DATA_BLOCK "DB_SDC_TS_PARAMETER_4"   // DB3707
{ S7_Optimized_Access := 'FALSE' }
AUTHOR : FFM
FAMILY : SDC
NAME : SECT_DEF
VERSION : 1.0
   VAR
      HEADER : Struct   // Struktur für Datenheader // nicht verschieben
         DB_NR : Int := 3707;   // DB Nummer
         MIN_NR_SEK : Int := 301;   // Niedrigste SEK Nummer im DB
         MAX_NR_SEK : Int := 400;   // Höchste SEK Nummer im DB
         START_DAT : Int := 20;   // Startadresse der SEK im DB
         LAENGE_SEK_DATA : Int := 260;   // Länge SEK Data
         ANZ_PROFIL : Int := 10;   // Number of Profiles
         OFFEST_PROFIL : Int := 40;   // Offestadresse der Profilparameter im TS-Parameterdatensatz
         LAENGE_PROFIL_DATA : Int := 22;   // Länge SEK Data
         Res160 : Int := 0;   // Reserve
         Res : Int := 0;   // Reserve
      END_STRUCT;
      TS : Array[301..400] of "UDT_SDC_TS_PARAMETER";
   END_VAR
BEGIN
   TS[301].ALLG.SEK_NEXT_1 := 0;
   TS[301].ALLG.SEK_NEXT_2 := 0;
   TS[301].ALLG.Spare[4] := 16#00;
   TS[301].ALLG.Spare[5] := 16#00;
   TS[301].ALLG.POS.Start_1 := 0;
   TS[301].ALLG.POS.End_1 := 0;
   TS[301].ALLG.POS.Start_2 := 0;
   TS[301].ALLG.POS.End_2 := 0;
   TS[301].ALLG.POS.Actionpoint_1 := 0;
   TS[301].ALLG.POS.Actionpoint_2 := 0;
   TS[301].ALLG.FLAGS.DIST_VAL[0] := TRUE;
   TS[301].ALLG.FLAGS.DIST_VAL[1] := FALSE;
   TS[301].ALLG.FLAGS.DIST_VAL[2] := FALSE;
   TS[301].ALLG.FLAGS.DIST_VAL[3] := FALSE;
   TS[301].ALLG.FLAGS.DIST_VAL[4] := FALSE;
   TS[301].ALLG.FLAGS.DIST_VAL[5] := FALSE;
   TS[301].ALLG.FLAGS.DIST_VAL[6] := FALSE;
   TS[301].ALLG.FLAGS.DIST_VAL[7] := FALSE;
   TS[301].ALLG.FLAGS.DIST_VAL[8] := FALSE;
   TS[301].ALLG.FLAGS.DIST_VAL[9] := FALSE;
   TS[301].ALLG.FLAGS.DIST_VAL[10] := FALSE;
   TS[301].ALLG.FLAGS.DIST_VAL[11] := FALSE;
   TS[301].ALLG.FLAGS.DIST_VAL[12] := FALSE;
   TS[301].ALLG.FLAGS.DIST_VAL[13] := FALSE;
   TS[301].ALLG.FLAGS.DIST_VAL[14] := FALSE;
   TS[301].ALLG.FLAGS.DIST_VAL[15] := FALSE;
   TS[301].ALLG.FLAGS.one_profile := FALSE;
   TS[301].ALLG.FLAGS.BLIND := FALSE;
   TS[301].ALLG.FLAGS.NO_DIST_CONT := FALSE;
   TS[301].ALLG.FLAGS.SYNCH_AREA := FALSE;
   TS[301].ALLG.FLAGS.bit24 := FALSE;
   TS[301].ALLG.FLAGS.bit25 := FALSE;
   TS[301].ALLG.FLAGS.bit26 := FALSE;
   TS[301].ALLG.FLAGS.bit27 := FALSE;
   TS[301].ALLG.FLAGS.EN_HOIST := FALSE;
   TS[301].ALLG.FLAGS.D_RESET_AFTER := FALSE;
   TS[301].ALLG.FLAGS.D_PULK := FALSE;
   TS[301].ALLG.FLAGS.bit33 := FALSE;
   TS[301].ALLG.FLAGS.bit34 := FALSE;
   TS[301].ALLG.FLAGS.bit35 := FALSE;
   TS[301].ALLG.FLAGS.bit36 := FALSE;
   TS[301].ALLG.FLAGS.Deutronic_ON := FALSE;
   TS[301].ALLG.Stop_Position := 0;
   TS[301].ALLG.Drive_speed_1 := 0;
   TS[301].ALLG.Drive_speed_2 := 0;
   TS[301].PROFIL[1].Hoist_Pos_start := 0;
   TS[301].PROFIL[1].Height := 2651;
   TS[301].PROFIL[1].Hoist_speed := 2000;
   TS[301].PROFIL[1].Hoist_offset_1 := 0;
   TS[301].PROFIL[1].Hoist_offset_2 := 0;
   TS[301].PROFIL[1].Hoist_offset_3 := 0;
   TS[301].PROFIL[1].Hoist_offset_4 := 0;
   TS[301].PROFIL[1].Hoist_Start_offset_1 := 0;
   TS[301].PROFIL[1].Hoist_Start_offset_2 := 0;
   TS[301].PROFIL[1].Hoist_Start_offset_3 := 0;
   TS[301].PROFIL[1].Hoist_Start_offset_4 := 0;
   TS[301].PROFIL[2].Hoist_Pos_start := 0;
   TS[301].PROFIL[2].Height := 2651;
   TS[301].PROFIL[2].Hoist_speed := 2000;
   TS[301].PROFIL[2].Hoist_offset_1 := 0;
   TS[301].PROFIL[2].Hoist_offset_2 := 0;
   TS[301].PROFIL[2].Hoist_offset_3 := 0;
   TS[301].PROFIL[2].Hoist_offset_4 := 0;
   TS[301].PROFIL[2].Hoist_Start_offset_1 := 0;
   TS[301].PROFIL[2].Hoist_Start_offset_2 := 0;
   TS[301].PROFIL[2].Hoist_Start_offset_3 := 0;
   TS[301].PROFIL[2].Hoist_Start_offset_4 := 0;
   TS[301].PROFIL[3].Hoist_Pos_start := 0;
   TS[301].PROFIL[3].Height := 2651;
   TS[301].PROFIL[3].Hoist_speed := 2000;
   TS[301].PROFIL[3].Hoist_offset_1 := 0;
   TS[301].PROFIL[3].Hoist_offset_2 := 0;
   TS[301].PROFIL[3].Hoist_offset_3 := 0;
   TS[301].PROFIL[3].Hoist_offset_4 := 0;
   TS[301].PROFIL[3].Hoist_Start_offset_1 := 0;
   TS[301].PROFIL[3].Hoist_Start_offset_2 := 0;
   TS[301].PROFIL[3].Hoist_Start_offset_3 := 0;
   TS[301].PROFIL[3].Hoist_Start_offset_4 := 0;
   TS[301].PROFIL[4].Hoist_Pos_start := 0;
   TS[301].PROFIL[4].Height := 2651;
   TS[301].PROFIL[4].Hoist_speed := 2000;
   TS[301].PROFIL[4].Hoist_offset_1 := 0;
   TS[301].PROFIL[4].Hoist_offset_2 := 0;
   TS[301].PROFIL[4].Hoist_offset_3 := 0;
   TS[301].PROFIL[4].Hoist_offset_4 := 0;
   TS[301].PROFIL[4].Hoist_Start_offset_1 := 0;
   TS[301].PROFIL[4].Hoist_Start_offset_2 := 0;
   TS[301].PROFIL[4].Hoist_Start_offset_3 := 0;
   TS[301].PROFIL[4].Hoist_Start_offset_4 := 0;
   TS[301].PROFIL[5].Hoist_Pos_start := 0;
   TS[301].PROFIL[5].Height := 2651;
   TS[301].PROFIL[5].Hoist_speed := 2000;
   TS[301].PROFIL[5].Hoist_offset_1 := 0;
   TS[301].PROFIL[5].Hoist_offset_2 := 0;
   TS[301].PROFIL[5].Hoist_offset_3 := 0;
   TS[301].PROFIL[5].Hoist_offset_4 := 0;
   TS[301].PROFIL[5].Hoist_Start_offset_1 := 0;
   TS[301].PROFIL[5].Hoist_Start_offset_2 := 0;
   TS[301].PROFIL[5].Hoist_Start_offset_3 := 0;
   TS[301].PROFIL[5].Hoist_Start_offset_4 := 0;
   TS[301].PROFIL[6].Hoist_Pos_start := 0;
   TS[301].PROFIL[6].Height := 2651;
   TS[301].PROFIL[6].Hoist_speed := 2000;
   TS[301].PROFIL[6].Hoist_offset_1 := 0;
   TS[301].PROFIL[6].Hoist_offset_2 := 0;
   TS[301].PROFIL[6].Hoist_offset_3 := 0;
   TS[301].PROFIL[6].Hoist_offset_4 := 0;
   TS[301].PROFIL[6].Hoist_Start_offset_1 := 0;
   TS[301].PROFIL[6].Hoist_Start_offset_2 := 0;
   TS[301].PROFIL[6].Hoist_Start_offset_3 := 0;
   TS[301].PROFIL[6].Hoist_Start_offset_4 := 0;
   TS[301].PROFIL[7].Hoist_Pos_start := 0;
   TS[301].PROFIL[7].Height := 2651;
   TS[301].PROFIL[7].Hoist_speed := 2000;
   TS[301].PROFIL[7].Hoist_offset_1 := 0;
   TS[301].PROFIL[7].Hoist_offset_2 := 0;
   TS[301].PROFIL[7].Hoist_offset_3 := 0;
   TS[301].PROFIL[7].Hoist_offset_4 := 0;
   TS[301].PROFIL[7].Hoist_Start_offset_1 := 0;
   TS[301].PROFIL[7].Hoist_Start_offset_2 := 0;
   TS[301].PROFIL[7].Hoist_Start_offset_3 := 0;
   TS[301].PROFIL[7].Hoist_Start_offset_4 := 0;
   TS[301].PROFIL[8].Hoist_Pos_start := 0;
   TS[301].PROFIL[8].Height := 2651;
   TS[301].PROFIL[8].Hoist_speed := 2000;
   TS[301].PROFIL[8].Hoist_offset_1 := 0;
   TS[301].PROFIL[8].Hoist_offset_2 := 0;
   TS[301].PROFIL[8].Hoist_offset_3 := 0;
   TS[301].PROFIL[8].Hoist_offset_4 := 0;
   TS[301].PROFIL[8].Hoist_Start_offset_1 := 0;
   TS[301].PROFIL[8].Hoist_Start_offset_2 := 0;
   TS[301].PROFIL[8].Hoist_Start_offset_3 := 0;
   TS[301].PROFIL[8].Hoist_Start_offset_4 := 0;
   TS[301].PROFIL[9].Hoist_Pos_start := 0;
   TS[301].PROFIL[9].Height := 2651;
   TS[301].PROFIL[9].Hoist_speed := 2000;
   TS[301].PROFIL[9].Hoist_offset_1 := 0;
   TS[301].PROFIL[9].Hoist_offset_2 := 0;
   TS[301].PROFIL[9].Hoist_offset_3 := 0;
   TS[301].PROFIL[9].Hoist_offset_4 := 0;
   TS[301].PROFIL[9].Hoist_Start_offset_1 := 0;
   TS[301].PROFIL[9].Hoist_Start_offset_2 := 0;
   TS[301].PROFIL[9].Hoist_Start_offset_3 := 0;
   TS[301].PROFIL[9].Hoist_Start_offset_4 := 0;
   TS[301].PROFIL[10].Hoist_Pos_start := 0;
   TS[301].PROFIL[10].Height := 2651;
   TS[301].PROFIL[10].Hoist_speed := 2000;
   TS[301].PROFIL[10].Hoist_offset_1 := 0;
   TS[301].PROFIL[10].Hoist_offset_2 := 0;
   TS[301].PROFIL[10].Hoist_offset_3 := 0;
   TS[301].PROFIL[10].Hoist_offset_4 := 0;
   TS[301].PROFIL[10].Hoist_Start_offset_1 := 0;
   TS[301].PROFIL[10].Hoist_Start_offset_2 := 0;
   TS[301].PROFIL[10].Hoist_Start_offset_3 := 0;
   TS[301].PROFIL[10].Hoist_Start_offset_4 := 0;
   TS[302].ALLG.SEK_NEXT_1 := 0;
   TS[302].ALLG.SEK_NEXT_2 := 0;
   TS[302].ALLG.Spare[4] := 16#00;
   TS[302].ALLG.Spare[5] := 16#00;
   TS[302].ALLG.POS.Start_1 := 0;
   TS[302].ALLG.POS.End_1 := 0;
   TS[302].ALLG.POS.Start_2 := 0;
   TS[302].ALLG.POS.End_2 := 0;
   TS[302].ALLG.POS.Actionpoint_1 := 0;
   TS[302].ALLG.POS.Actionpoint_2 := 0;
   TS[302].ALLG.FLAGS.DIST_VAL[0] := TRUE;
   TS[302].ALLG.FLAGS.DIST_VAL[1] := FALSE;
   TS[302].ALLG.FLAGS.DIST_VAL[2] := FALSE;
   TS[302].ALLG.FLAGS.DIST_VAL[3] := FALSE;
   TS[302].ALLG.FLAGS.DIST_VAL[4] := FALSE;
   TS[302].ALLG.FLAGS.DIST_VAL[5] := FALSE;
   TS[302].ALLG.FLAGS.DIST_VAL[6] := FALSE;
   TS[302].ALLG.FLAGS.DIST_VAL[7] := FALSE;
   TS[302].ALLG.FLAGS.DIST_VAL[8] := FALSE;
   TS[302].ALLG.FLAGS.DIST_VAL[9] := FALSE;
   TS[302].ALLG.FLAGS.DIST_VAL[10] := FALSE;
   TS[302].ALLG.FLAGS.DIST_VAL[11] := FALSE;
   TS[302].ALLG.FLAGS.DIST_VAL[12] := FALSE;
   TS[302].ALLG.FLAGS.DIST_VAL[13] := FALSE;
   TS[302].ALLG.FLAGS.DIST_VAL[14] := FALSE;
   TS[302].ALLG.FLAGS.DIST_VAL[15] := FALSE;
   TS[302].ALLG.FLAGS.one_profile := FALSE;
   TS[302].ALLG.FLAGS.BLIND := FALSE;
   TS[302].ALLG.FLAGS.NO_DIST_CONT := FALSE;
   TS[302].ALLG.FLAGS.SYNCH_AREA := FALSE;
   TS[302].ALLG.FLAGS.bit24 := FALSE;
   TS[302].ALLG.FLAGS.bit25 := FALSE;
   TS[302].ALLG.FLAGS.bit26 := FALSE;
   TS[302].ALLG.FLAGS.bit27 := FALSE;
   TS[302].ALLG.FLAGS.EN_HOIST := FALSE;
   TS[302].ALLG.FLAGS.D_RESET_AFTER := FALSE;
   TS[302].ALLG.FLAGS.D_PULK := FALSE;
   TS[302].ALLG.FLAGS.bit33 := FALSE;
   TS[302].ALLG.FLAGS.bit34 := FALSE;
   TS[302].ALLG.FLAGS.bit35 := FALSE;
   TS[302].ALLG.FLAGS.bit36 := FALSE;
   TS[302].ALLG.FLAGS.Deutronic_ON := FALSE;
   TS[302].ALLG.Stop_Position := 0;
   TS[302].ALLG.Drive_speed_1 := 0;
   TS[302].ALLG.Drive_speed_2 := 0;
   // 15300 more start values not shown
END_DATA_BLOCK

DATA_BLOCK "DB_SDC_TS_PARAMETER_5"   // DB3708
{ S7_Optimized_Access := 'FALSE' }
AUTHOR : FFM
FAMILY : SDC
NAME : SECT_DEF
VERSION : 1.0
   VAR
      HEADER : Struct   // Struktur für Datenheader // nicht verschieben
         DB_NR : Int := 3708;   // DB Nummer
         MIN_NR_SEK : Int := 401;   // Niedrigste SEK Nummer im DB
         MAX_NR_SEK : Int := 500;   // Höchste SEK Nummer im DB
         START_DAT : Int := 20;   // Startadresse der SEK im DB
         LAENGE_SEK_DATA : Int := 260;   // Länge SEK Data
         ANZ_PROFIL : Int := 10;   // Number of Profiles
         OFFEST_PROFIL : Int := 40;   // Offestadresse der Profilparameter im TS-Parameterdatensatz
         LAENGE_PROFIL_DATA : Int := 22;   // Länge SEK Data
         Res160 : Int := 0;   // Reserve
         Res : Int := 0;   // Reserve
      END_STRUCT;
      TS : Array[401..500] of "UDT_SDC_TS_PARAMETER";
   END_VAR
BEGIN
   TS[401].ALLG.SEK_NEXT_1 := 0;
   TS[401].ALLG.SEK_NEXT_2 := 0;
   TS[401].ALLG.Spare[4] := 16#00;
   TS[401].ALLG.Spare[5] := 16#00;
   TS[401].ALLG.POS.Start_1 := 1159500;
   TS[401].ALLG.POS.End_1 := 1165999;
   TS[401].ALLG.POS.Start_2 := 0;
   TS[401].ALLG.POS.End_2 := 0;
   TS[401].ALLG.POS.Actionpoint_1 := 0;
   TS[401].ALLG.POS.Actionpoint_2 := 0;
   TS[401].ALLG.FLAGS.DIST_VAL[0] := FALSE;
   TS[401].ALLG.FLAGS.DIST_VAL[1] := FALSE;
   TS[401].ALLG.FLAGS.DIST_VAL[2] := FALSE;
   TS[401].ALLG.FLAGS.DIST_VAL[3] := FALSE;
   TS[401].ALLG.FLAGS.DIST_VAL[4] := FALSE;
   TS[401].ALLG.FLAGS.DIST_VAL[5] := FALSE;
   TS[401].ALLG.FLAGS.DIST_VAL[6] := FALSE;
   TS[401].ALLG.FLAGS.DIST_VAL[7] := FALSE;
   TS[401].ALLG.FLAGS.DIST_VAL[8] := FALSE;
   TS[401].ALLG.FLAGS.DIST_VAL[9] := TRUE;
   TS[401].ALLG.FLAGS.DIST_VAL[10] := FALSE;
   TS[401].ALLG.FLAGS.DIST_VAL[11] := FALSE;
   TS[401].ALLG.FLAGS.DIST_VAL[12] := FALSE;
   TS[401].ALLG.FLAGS.DIST_VAL[13] := FALSE;
   TS[401].ALLG.FLAGS.DIST_VAL[14] := FALSE;
   TS[401].ALLG.FLAGS.DIST_VAL[15] := FALSE;
   TS[401].ALLG.FLAGS.one_profile := FALSE;
   TS[401].ALLG.FLAGS.BLIND := FALSE;
   TS[401].ALLG.FLAGS.NO_DIST_CONT := FALSE;
   TS[401].ALLG.FLAGS.SYNCH_AREA := FALSE;
   TS[401].ALLG.FLAGS.bit24 := FALSE;
   TS[401].ALLG.FLAGS.bit25 := FALSE;
   TS[401].ALLG.FLAGS.bit26 := FALSE;
   TS[401].ALLG.FLAGS.bit27 := FALSE;
   TS[401].ALLG.FLAGS.EN_HOIST := FALSE;
   TS[401].ALLG.FLAGS.D_RESET_AFTER := FALSE;
   TS[401].ALLG.FLAGS.D_PULK := FALSE;
   TS[401].ALLG.FLAGS.bit33 := FALSE;
   TS[401].ALLG.FLAGS.bit34 := FALSE;
   TS[401].ALLG.FLAGS.bit35 := FALSE;
   TS[401].ALLG.FLAGS.bit36 := FALSE;
   TS[401].ALLG.FLAGS.Deutronic_ON := FALSE;
   TS[401].ALLG.Stop_Position := 5800;
   TS[401].ALLG.Drive_speed_1 := 15000;
   TS[401].ALLG.Drive_speed_2 := 6000;
   TS[401].PROFIL[1].Hoist_Pos_start := 0;
   TS[401].PROFIL[1].Height := 3890;
   TS[401].PROFIL[1].Hoist_speed := 2000;
   TS[401].PROFIL[1].Hoist_offset_1 := 0;
   TS[401].PROFIL[1].Hoist_offset_2 := 0;
   TS[401].PROFIL[1].Hoist_offset_3 := 0;
   TS[401].PROFIL[1].Hoist_offset_4 := 0;
   TS[401].PROFIL[1].Hoist_Start_offset_1 := 0;
   TS[401].PROFIL[1].Hoist_Start_offset_2 := 0;
   TS[401].PROFIL[1].Hoist_Start_offset_3 := 0;
   TS[401].PROFIL[1].Hoist_Start_offset_4 := 0;
   TS[401].PROFIL[2].Hoist_Pos_start := 0;
   TS[401].PROFIL[2].Height := 3890;
   TS[401].PROFIL[2].Hoist_speed := 2000;
   TS[401].PROFIL[2].Hoist_offset_1 := 0;
   TS[401].PROFIL[2].Hoist_offset_2 := 0;
   TS[401].PROFIL[2].Hoist_offset_3 := 0;
   TS[401].PROFIL[2].Hoist_offset_4 := 0;
   TS[401].PROFIL[2].Hoist_Start_offset_1 := 0;
   TS[401].PROFIL[2].Hoist_Start_offset_2 := 0;
   TS[401].PROFIL[2].Hoist_Start_offset_3 := 0;
   TS[401].PROFIL[2].Hoist_Start_offset_4 := 0;
   TS[401].PROFIL[3].Hoist_Pos_start := 0;
   TS[401].PROFIL[3].Height := 3890;
   TS[401].PROFIL[3].Hoist_speed := 2000;
   TS[401].PROFIL[3].Hoist_offset_1 := 0;
   TS[401].PROFIL[3].Hoist_offset_2 := 0;
   TS[401].PROFIL[3].Hoist_offset_3 := 0;
   TS[401].PROFIL[3].Hoist_offset_4 := 0;
   TS[401].PROFIL[3].Hoist_Start_offset_1 := 0;
   TS[401].PROFIL[3].Hoist_Start_offset_2 := 0;
   TS[401].PROFIL[3].Hoist_Start_offset_3 := 0;
   TS[401].PROFIL[3].Hoist_Start_offset_4 := 0;
   TS[401].PROFIL[4].Hoist_Pos_start := 0;
   TS[401].PROFIL[4].Height := 3890;
   TS[401].PROFIL[4].Hoist_speed := 2000;
   TS[401].PROFIL[4].Hoist_offset_1 := 0;
   TS[401].PROFIL[4].Hoist_offset_2 := 0;
   TS[401].PROFIL[4].Hoist_offset_3 := 0;
   TS[401].PROFIL[4].Hoist_offset_4 := 0;
   TS[401].PROFIL[4].Hoist_Start_offset_1 := 0;
   TS[401].PROFIL[4].Hoist_Start_offset_2 := 0;
   TS[401].PROFIL[4].Hoist_Start_offset_3 := 0;
   TS[401].PROFIL[4].Hoist_Start_offset_4 := 0;
   TS[401].PROFIL[5].Hoist_Pos_start := 0;
   TS[401].PROFIL[5].Height := 3890;
   TS[401].PROFIL[5].Hoist_speed := 2000;
   TS[401].PROFIL[5].Hoist_offset_1 := 0;
   TS[401].PROFIL[5].Hoist_offset_2 := 0;
   TS[401].PROFIL[5].Hoist_offset_3 := 0;
   TS[401].PROFIL[5].Hoist_offset_4 := 0;
   TS[401].PROFIL[5].Hoist_Start_offset_1 := 0;
   TS[401].PROFIL[5].Hoist_Start_offset_2 := 0;
   TS[401].PROFIL[5].Hoist_Start_offset_3 := 0;
   TS[401].PROFIL[5].Hoist_Start_offset_4 := 0;
   TS[401].PROFIL[6].Hoist_Pos_start := 0;
   TS[401].PROFIL[6].Height := 3890;
   TS[401].PROFIL[6].Hoist_speed := 2000;
   TS[401].PROFIL[6].Hoist_offset_1 := 0;
   TS[401].PROFIL[6].Hoist_offset_2 := 0;
   TS[401].PROFIL[6].Hoist_offset_3 := 0;
   TS[401].PROFIL[6].Hoist_offset_4 := 0;
   TS[401].PROFIL[6].Hoist_Start_offset_1 := 0;
   TS[401].PROFIL[6].Hoist_Start_offset_2 := 0;
   TS[401].PROFIL[6].Hoist_Start_offset_3 := 0;
   TS[401].PROFIL[6].Hoist_Start_offset_4 := 0;
   TS[401].PROFIL[7].Hoist_Pos_start := 0;
   TS[401].PROFIL[7].Height := 3890;
   TS[401].PROFIL[7].Hoist_speed := 2000;
   TS[401].PROFIL[7].Hoist_offset_1 := 0;
   TS[401].PROFIL[7].Hoist_offset_2 := 0;
   TS[401].PROFIL[7].Hoist_offset_3 := 0;
   TS[401].PROFIL[7].Hoist_offset_4 := 0;
   TS[401].PROFIL[7].Hoist_Start_offset_1 := 0;
   TS[401].PROFIL[7].Hoist_Start_offset_2 := 0;
   TS[401].PROFIL[7].Hoist_Start_offset_3 := 0;
   TS[401].PROFIL[7].Hoist_Start_offset_4 := 0;
   TS[401].PROFIL[8].Hoist_Pos_start := 0;
   TS[401].PROFIL[8].Height := 3890;
   TS[401].PROFIL[8].Hoist_speed := 2000;
   TS[401].PROFIL[8].Hoist_offset_1 := 0;
   TS[401].PROFIL[8].Hoist_offset_2 := 0;
   TS[401].PROFIL[8].Hoist_offset_3 := 0;
   TS[401].PROFIL[8].Hoist_offset_4 := 0;
   TS[401].PROFIL[8].Hoist_Start_offset_1 := 0;
   TS[401].PROFIL[8].Hoist_Start_offset_2 := 0;
   TS[401].PROFIL[8].Hoist_Start_offset_3 := 0;
   TS[401].PROFIL[8].Hoist_Start_offset_4 := 0;
   TS[401].PROFIL[9].Hoist_Pos_start := 0;
   TS[401].PROFIL[9].Height := 3890;
   TS[401].PROFIL[9].Hoist_speed := 2000;
   TS[401].PROFIL[9].Hoist_offset_1 := 0;
   TS[401].PROFIL[9].Hoist_offset_2 := 0;
   TS[401].PROFIL[9].Hoist_offset_3 := 0;
   TS[401].PROFIL[9].Hoist_offset_4 := 0;
   TS[401].PROFIL[9].Hoist_Start_offset_1 := 0;
   TS[401].PROFIL[9].Hoist_Start_offset_2 := 0;
   TS[401].PROFIL[9].Hoist_Start_offset_3 := 0;
   TS[401].PROFIL[9].Hoist_Start_offset_4 := 0;
   TS[401].PROFIL[10].Hoist_Pos_start := 0;
   TS[401].PROFIL[10].Height := 3890;
   TS[401].PROFIL[10].Hoist_speed := 2000;
   TS[401].PROFIL[10].Hoist_offset_1 := 0;
   TS[401].PROFIL[10].Hoist_offset_2 := 0;
   TS[401].PROFIL[10].Hoist_offset_3 := 0;
   TS[401].PROFIL[10].Hoist_offset_4 := 0;
   TS[401].PROFIL[10].Hoist_Start_offset_1 := 0;
   TS[401].PROFIL[10].Hoist_Start_offset_2 := 0;
   TS[401].PROFIL[10].Hoist_Start_offset_3 := 0;
   TS[401].PROFIL[10].Hoist_Start_offset_4 := 0;
   TS[402].ALLG.SEK_NEXT_1 := 0;
   TS[402].ALLG.SEK_NEXT_2 := 0;
   TS[402].ALLG.Spare[4] := 16#00;
   TS[402].ALLG.Spare[5] := 16#00;
   TS[402].ALLG.POS.Start_1 := 1166000;
   TS[402].ALLG.POS.End_1 := 1172199;
   TS[402].ALLG.POS.Start_2 := 0;
   TS[402].ALLG.POS.End_2 := 0;
   TS[402].ALLG.POS.Actionpoint_1 := 0;
   TS[402].ALLG.POS.Actionpoint_2 := 0;
   TS[402].ALLG.FLAGS.DIST_VAL[0] := FALSE;
   TS[402].ALLG.FLAGS.DIST_VAL[1] := FALSE;
   TS[402].ALLG.FLAGS.DIST_VAL[2] := FALSE;
   TS[402].ALLG.FLAGS.DIST_VAL[3] := FALSE;
   TS[402].ALLG.FLAGS.DIST_VAL[4] := FALSE;
   TS[402].ALLG.FLAGS.DIST_VAL[5] := TRUE;
   TS[402].ALLG.FLAGS.DIST_VAL[6] := FALSE;
   TS[402].ALLG.FLAGS.DIST_VAL[7] := FALSE;
   TS[402].ALLG.FLAGS.DIST_VAL[8] := FALSE;
   TS[402].ALLG.FLAGS.DIST_VAL[9] := FALSE;
   TS[402].ALLG.FLAGS.DIST_VAL[10] := FALSE;
   TS[402].ALLG.FLAGS.DIST_VAL[11] := FALSE;
   TS[402].ALLG.FLAGS.DIST_VAL[12] := FALSE;
   TS[402].ALLG.FLAGS.DIST_VAL[13] := FALSE;
   TS[402].ALLG.FLAGS.DIST_VAL[14] := FALSE;
   TS[402].ALLG.FLAGS.DIST_VAL[15] := FALSE;
   TS[402].ALLG.FLAGS.one_profile := FALSE;
   TS[402].ALLG.FLAGS.BLIND := FALSE;
   TS[402].ALLG.FLAGS.NO_DIST_CONT := FALSE;
   TS[402].ALLG.FLAGS.SYNCH_AREA := FALSE;
   TS[402].ALLG.FLAGS.bit24 := FALSE;
   TS[402].ALLG.FLAGS.bit25 := FALSE;
   TS[402].ALLG.FLAGS.bit26 := FALSE;
   TS[402].ALLG.FLAGS.bit27 := FALSE;
   TS[402].ALLG.FLAGS.EN_HOIST := FALSE;
   TS[402].ALLG.FLAGS.D_RESET_AFTER := FALSE;
   TS[402].ALLG.FLAGS.D_PULK := FALSE;
   TS[402].ALLG.FLAGS.bit33 := FALSE;
   TS[402].ALLG.FLAGS.bit34 := FALSE;
   TS[402].ALLG.FLAGS.bit35 := FALSE;
   TS[402].ALLG.FLAGS.bit36 := FALSE;
   TS[402].ALLG.FLAGS.Deutronic_ON := FALSE;
   TS[402].ALLG.Stop_Position := 5800;
   TS[402].ALLG.Drive_speed_1 := 15000;
   TS[402].ALLG.Drive_speed_2 := 6000;
   // 15300 more start values not shown
END_DATA_BLOCK

DATA_BLOCK "DB_SDC_TS_PARAMETER_6"   // DB3709
{ S7_Optimized_Access := 'FALSE' }
AUTHOR : FFM
FAMILY : SDC
NAME : SECT_DEF
VERSION : 1.0
   VAR
      HEADER : Struct   // Struktur für Datenheader // nicht verschieben
         DB_NR : Int := 3709;   // DB Nummer
         MIN_NR_SEK : Int := 501;   // Niedrigste SEK Nummer im DB
         MAX_NR_SEK : Int := 600;   // Höchste SEK Nummer im DB
         START_DAT : Int := 20;   // Startadresse der SEK im DB
         LAENGE_SEK_DATA : Int := 260;   // Länge SEK Data
         ANZ_PROFIL : Int := 10;   // Number of Profiles
         OFFEST_PROFIL : Int := 40;   // Offestadresse der Profilparameter im TS-Parameterdatensatz
         LAENGE_PROFIL_DATA : Int := 22;   // Länge SEK Data
         Res160 : Int := 0;   // Reserve
         Res : Int := 0;   // Reserve
      END_STRUCT;
      TS : Array[501..600] of "UDT_SDC_TS_PARAMETER";
   END_VAR
BEGIN
   TS[501].ALLG.SEK_NEXT_1 := 0;
   TS[501].ALLG.SEK_NEXT_2 := 0;
   TS[501].ALLG.Spare[4] := 16#00;
   TS[501].ALLG.Spare[5] := 16#00;
   TS[501].ALLG.POS.Start_1 := 1639750;
   TS[501].ALLG.POS.End_1 := 1646749;
   TS[501].ALLG.POS.Start_2 := 0;
   TS[501].ALLG.POS.End_2 := 0;
   TS[501].ALLG.POS.Actionpoint_1 := 0;
   TS[501].ALLG.POS.Actionpoint_2 := 0;
   TS[501].ALLG.FLAGS.DIST_VAL[0] := FALSE;
   TS[501].ALLG.FLAGS.DIST_VAL[1] := FALSE;
   TS[501].ALLG.FLAGS.DIST_VAL[2] := FALSE;
   TS[501].ALLG.FLAGS.DIST_VAL[3] := FALSE;
   TS[501].ALLG.FLAGS.DIST_VAL[4] := FALSE;
   TS[501].ALLG.FLAGS.DIST_VAL[5] := FALSE;
   TS[501].ALLG.FLAGS.DIST_VAL[6] := FALSE;
   TS[501].ALLG.FLAGS.DIST_VAL[7] := FALSE;
   TS[501].ALLG.FLAGS.DIST_VAL[8] := FALSE;
   TS[501].ALLG.FLAGS.DIST_VAL[9] := TRUE;
   TS[501].ALLG.FLAGS.DIST_VAL[10] := FALSE;
   TS[501].ALLG.FLAGS.DIST_VAL[11] := FALSE;
   TS[501].ALLG.FLAGS.DIST_VAL[12] := FALSE;
   TS[501].ALLG.FLAGS.DIST_VAL[13] := FALSE;
   TS[501].ALLG.FLAGS.DIST_VAL[14] := FALSE;
   TS[501].ALLG.FLAGS.DIST_VAL[15] := FALSE;
   TS[501].ALLG.FLAGS.one_profile := FALSE;
   TS[501].ALLG.FLAGS.BLIND := FALSE;
   TS[501].ALLG.FLAGS.NO_DIST_CONT := FALSE;
   TS[501].ALLG.FLAGS.SYNCH_AREA := FALSE;
   TS[501].ALLG.FLAGS.bit24 := FALSE;
   TS[501].ALLG.FLAGS.bit25 := FALSE;
   TS[501].ALLG.FLAGS.bit26 := FALSE;
   TS[501].ALLG.FLAGS.bit27 := FALSE;
   TS[501].ALLG.FLAGS.EN_HOIST := FALSE;
   TS[501].ALLG.FLAGS.D_RESET_AFTER := FALSE;
   TS[501].ALLG.FLAGS.D_PULK := FALSE;
   TS[501].ALLG.FLAGS.bit33 := FALSE;
   TS[501].ALLG.FLAGS.bit34 := FALSE;
   TS[501].ALLG.FLAGS.bit35 := FALSE;
   TS[501].ALLG.FLAGS.bit36 := FALSE;
   TS[501].ALLG.FLAGS.Deutronic_ON := FALSE;
   TS[501].ALLG.Stop_Position := 6500;
   TS[501].ALLG.Drive_speed_1 := 15000;
   TS[501].ALLG.Drive_speed_2 := 6000;
   TS[501].PROFIL[1].Hoist_Pos_start := 0;
   TS[501].PROFIL[1].Height := 3890;
   TS[501].PROFIL[1].Hoist_speed := 2000;
   TS[501].PROFIL[1].Hoist_offset_1 := 0;
   TS[501].PROFIL[1].Hoist_offset_2 := 0;
   TS[501].PROFIL[1].Hoist_offset_3 := 0;
   TS[501].PROFIL[1].Hoist_offset_4 := 0;
   TS[501].PROFIL[1].Hoist_Start_offset_1 := 0;
   TS[501].PROFIL[1].Hoist_Start_offset_2 := 0;
   TS[501].PROFIL[1].Hoist_Start_offset_3 := 0;
   TS[501].PROFIL[1].Hoist_Start_offset_4 := 0;
   TS[501].PROFIL[2].Hoist_Pos_start := 0;
   TS[501].PROFIL[2].Height := 3890;
   TS[501].PROFIL[2].Hoist_speed := 2000;
   TS[501].PROFIL[2].Hoist_offset_1 := 0;
   TS[501].PROFIL[2].Hoist_offset_2 := 0;
   TS[501].PROFIL[2].Hoist_offset_3 := 0;
   TS[501].PROFIL[2].Hoist_offset_4 := 0;
   TS[501].PROFIL[2].Hoist_Start_offset_1 := 0;
   TS[501].PROFIL[2].Hoist_Start_offset_2 := 0;
   TS[501].PROFIL[2].Hoist_Start_offset_3 := 0;
   TS[501].PROFIL[2].Hoist_Start_offset_4 := 0;
   TS[501].PROFIL[3].Hoist_Pos_start := 0;
   TS[501].PROFIL[3].Height := 3890;
   TS[501].PROFIL[3].Hoist_speed := 2000;
   TS[501].PROFIL[3].Hoist_offset_1 := 0;
   TS[501].PROFIL[3].Hoist_offset_2 := 0;
   TS[501].PROFIL[3].Hoist_offset_3 := 0;
   TS[501].PROFIL[3].Hoist_offset_4 := 0;
   TS[501].PROFIL[3].Hoist_Start_offset_1 := 0;
   TS[501].PROFIL[3].Hoist_Start_offset_2 := 0;
   TS[501].PROFIL[3].Hoist_Start_offset_3 := 0;
   TS[501].PROFIL[3].Hoist_Start_offset_4 := 0;
   TS[501].PROFIL[4].Hoist_Pos_start := 0;
   TS[501].PROFIL[4].Height := 3890;
   TS[501].PROFIL[4].Hoist_speed := 2000;
   TS[501].PROFIL[4].Hoist_offset_1 := 0;
   TS[501].PROFIL[4].Hoist_offset_2 := 0;
   TS[501].PROFIL[4].Hoist_offset_3 := 0;
   TS[501].PROFIL[4].Hoist_offset_4 := 0;
   TS[501].PROFIL[4].Hoist_Start_offset_1 := 0;
   TS[501].PROFIL[4].Hoist_Start_offset_2 := 0;
   TS[501].PROFIL[4].Hoist_Start_offset_3 := 0;
   TS[501].PROFIL[4].Hoist_Start_offset_4 := 0;
   TS[501].PROFIL[5].Hoist_Pos_start := 0;
   TS[501].PROFIL[5].Height := 3890;
   TS[501].PROFIL[5].Hoist_speed := 2000;
   TS[501].PROFIL[5].Hoist_offset_1 := 0;
   TS[501].PROFIL[5].Hoist_offset_2 := 0;
   TS[501].PROFIL[5].Hoist_offset_3 := 0;
   TS[501].PROFIL[5].Hoist_offset_4 := 0;
   TS[501].PROFIL[5].Hoist_Start_offset_1 := 0;
   TS[501].PROFIL[5].Hoist_Start_offset_2 := 0;
   TS[501].PROFIL[5].Hoist_Start_offset_3 := 0;
   TS[501].PROFIL[5].Hoist_Start_offset_4 := 0;
   TS[501].PROFIL[6].Hoist_Pos_start := 0;
   TS[501].PROFIL[6].Height := 3890;
   TS[501].PROFIL[6].Hoist_speed := 2000;
   TS[501].PROFIL[6].Hoist_offset_1 := 0;
   TS[501].PROFIL[6].Hoist_offset_2 := 0;
   TS[501].PROFIL[6].Hoist_offset_3 := 0;
   TS[501].PROFIL[6].Hoist_offset_4 := 0;
   TS[501].PROFIL[6].Hoist_Start_offset_1 := 0;
   TS[501].PROFIL[6].Hoist_Start_offset_2 := 0;
   TS[501].PROFIL[6].Hoist_Start_offset_3 := 0;
   TS[501].PROFIL[6].Hoist_Start_offset_4 := 0;
   TS[501].PROFIL[7].Hoist_Pos_start := 0;
   TS[501].PROFIL[7].Height := 3890;
   TS[501].PROFIL[7].Hoist_speed := 2000;
   TS[501].PROFIL[7].Hoist_offset_1 := 0;
   TS[501].PROFIL[7].Hoist_offset_2 := 0;
   TS[501].PROFIL[7].Hoist_offset_3 := 0;
   TS[501].PROFIL[7].Hoist_offset_4 := 0;
   TS[501].PROFIL[7].Hoist_Start_offset_1 := 0;
   TS[501].PROFIL[7].Hoist_Start_offset_2 := 0;
   TS[501].PROFIL[7].Hoist_Start_offset_3 := 0;
   TS[501].PROFIL[7].Hoist_Start_offset_4 := 0;
   TS[501].PROFIL[8].Hoist_Pos_start := 0;
   TS[501].PROFIL[8].Height := 3890;
   TS[501].PROFIL[8].Hoist_speed := 2000;
   TS[501].PROFIL[8].Hoist_offset_1 := 0;
   TS[501].PROFIL[8].Hoist_offset_2 := 0;
   TS[501].PROFIL[8].Hoist_offset_3 := 0;
   TS[501].PROFIL[8].Hoist_offset_4 := 0;
   TS[501].PROFIL[8].Hoist_Start_offset_1 := 0;
   TS[501].PROFIL[8].Hoist_Start_offset_2 := 0;
   TS[501].PROFIL[8].Hoist_Start_offset_3 := 0;
   TS[501].PROFIL[8].Hoist_Start_offset_4 := 0;
   TS[501].PROFIL[9].Hoist_Pos_start := 0;
   TS[501].PROFIL[9].Height := 3890;
   TS[501].PROFIL[9].Hoist_speed := 2000;
   TS[501].PROFIL[9].Hoist_offset_1 := 0;
   TS[501].PROFIL[9].Hoist_offset_2 := 0;
   TS[501].PROFIL[9].Hoist_offset_3 := 0;
   TS[501].PROFIL[9].Hoist_offset_4 := 0;
   TS[501].PROFIL[9].Hoist_Start_offset_1 := 0;
   TS[501].PROFIL[9].Hoist_Start_offset_2 := 0;
   TS[501].PROFIL[9].Hoist_Start_offset_3 := 0;
   TS[501].PROFIL[9].Hoist_Start_offset_4 := 0;
   TS[501].PROFIL[10].Hoist_Pos_start := 0;
   TS[501].PROFIL[10].Height := 3890;
   TS[501].PROFIL[10].Hoist_speed := 2000;
   TS[501].PROFIL[10].Hoist_offset_1 := 0;
   TS[501].PROFIL[10].Hoist_offset_2 := 0;
   TS[501].PROFIL[10].Hoist_offset_3 := 0;
   TS[501].PROFIL[10].Hoist_offset_4 := 0;
   TS[501].PROFIL[10].Hoist_Start_offset_1 := 0;
   TS[501].PROFIL[10].Hoist_Start_offset_2 := 0;
   TS[501].PROFIL[10].Hoist_Start_offset_3 := 0;
   TS[501].PROFIL[10].Hoist_Start_offset_4 := 0;
   TS[502].ALLG.SEK_NEXT_1 := 0;
   TS[502].ALLG.SEK_NEXT_2 := 0;
   TS[502].ALLG.Spare[4] := 16#00;
   TS[502].ALLG.Spare[5] := 16#00;
   TS[502].ALLG.POS.Start_1 := 1646750;
   TS[502].ALLG.POS.End_1 := 1653749;
   TS[502].ALLG.POS.Start_2 := 0;
   TS[502].ALLG.POS.End_2 := 0;
   TS[502].ALLG.POS.Actionpoint_1 := 0;
   TS[502].ALLG.POS.Actionpoint_2 := 0;
   TS[502].ALLG.FLAGS.DIST_VAL[0] := FALSE;
   TS[502].ALLG.FLAGS.DIST_VAL[1] := FALSE;
   TS[502].ALLG.FLAGS.DIST_VAL[2] := FALSE;
   TS[502].ALLG.FLAGS.DIST_VAL[3] := FALSE;
   TS[502].ALLG.FLAGS.DIST_VAL[4] := FALSE;
   TS[502].ALLG.FLAGS.DIST_VAL[5] := FALSE;
   TS[502].ALLG.FLAGS.DIST_VAL[6] := FALSE;
   TS[502].ALLG.FLAGS.DIST_VAL[7] := FALSE;
   TS[502].ALLG.FLAGS.DIST_VAL[8] := FALSE;
   TS[502].ALLG.FLAGS.DIST_VAL[9] := TRUE;
   TS[502].ALLG.FLAGS.DIST_VAL[10] := FALSE;
   TS[502].ALLG.FLAGS.DIST_VAL[11] := FALSE;
   TS[502].ALLG.FLAGS.DIST_VAL[12] := FALSE;
   TS[502].ALLG.FLAGS.DIST_VAL[13] := FALSE;
   TS[502].ALLG.FLAGS.DIST_VAL[14] := FALSE;
   TS[502].ALLG.FLAGS.DIST_VAL[15] := FALSE;
   TS[502].ALLG.FLAGS.one_profile := FALSE;
   TS[502].ALLG.FLAGS.BLIND := FALSE;
   TS[502].ALLG.FLAGS.NO_DIST_CONT := FALSE;
   TS[502].ALLG.FLAGS.SYNCH_AREA := FALSE;
   TS[502].ALLG.FLAGS.bit24 := FALSE;
   TS[502].ALLG.FLAGS.bit25 := FALSE;
   TS[502].ALLG.FLAGS.bit26 := FALSE;
   TS[502].ALLG.FLAGS.bit27 := FALSE;
   TS[502].ALLG.FLAGS.EN_HOIST := FALSE;
   TS[502].ALLG.FLAGS.D_RESET_AFTER := FALSE;
   TS[502].ALLG.FLAGS.D_PULK := FALSE;
   TS[502].ALLG.FLAGS.bit33 := FALSE;
   TS[502].ALLG.FLAGS.bit34 := FALSE;
   TS[502].ALLG.FLAGS.bit35 := FALSE;
   TS[502].ALLG.FLAGS.bit36 := FALSE;
   TS[502].ALLG.FLAGS.Deutronic_ON := FALSE;
   TS[502].ALLG.Stop_Position := 6400;
   TS[502].ALLG.Drive_speed_1 := 15000;
   TS[502].ALLG.Drive_speed_2 := 6000;
   // 15300 more start values not shown
END_DATA_BLOCK

DATA_BLOCK "DB_SDC_EMS_1"   // DB3714
{ S7_Optimized_Access := 'FALSE' }
VERSION : 0.1
   VAR
      HEADER : Struct
         DB_NR : Int := 3714;
         MIN_NR_EMS : Int := 1;
         MAX_NR_EMS : Int := 200;
         START_EMS : Int := 20;
         LAENGE_EMS : Int := 260;
         OFFSET_EMS_SEK_STAT : Int := 164;
         LAENGE_EMS_SEK_STAT : Int := 34;
         OFFSET_EMS_FKT : Int := 216;
         Res160 : Int := 0;
         Load : Bool := TRUE;
      END_STRUCT;
   END_VAR
BEGIN
END_DATA_BLOCK

DATA_BLOCK "DB_SDC_TS_IF_COMMAND"   // DB3716
{ S7_Optimized_Access := 'FALSE' }
AUTHOR : FFM
FAMILY : SDC
NAME : SECT_IF
VERSION : 0.1
   VAR
      HEADER : Struct   // Struktur für Datenheader // nicht verschieben
         DB_NR : Int := 3716;   // DB Nummer
         MIN_NR_SEK : Int := 1;   // Niedrigste SEK Nummer im DB
         MAX_NR_SEK : Int := 600;   // Höchste SEK Nummer im DB
         START_DAT : Int := 20;   // Startadresse der SEK im DB
         LAENGE_SEK_DATA : Int := 18;   // Länge SEK Data
         LAENGE_VAL_DATA : Int := 8;   // Länge Value Data
         LAENGE_BIT_DATA : Int := 6;   // Länge Bit Data
         LAENGE_FKT : Int := 4;   // Länge Funktion
         Res16 : Int;   // Reserve
         Res18 : Int;   // Reserve
      END_STRUCT;
      SEK : Array[1..600] of "UDT_SDC_EMS_TS_COM";   // Komando für Sektion
   END_VAR
BEGIN
END_DATA_BLOCK

DATA_BLOCK "DB_SDC_TS_IF_COMMAND_2"   // DB3717
{ S7_Optimized_Access := 'FALSE' }
AUTHOR : FFM
FAMILY : SDC
NAME : SECT_IF
VERSION : 0.1
   VAR
      HEADER : Struct   // Struktur für Datenheader // nicht verschieben
         DB_NR : Int := 3717;   // DB Nummer
         MIN_NR_SEK : Int := 601;   // Niedrigste SEK Nummer im DB
         MAX_NR_SEK : Int := 1000;   // Höchste SEK Nummer im DB
         START_DAT : Int := 20;   // Startadresse der SEK im DB
         LAENGE_SEK_DATA : Int := 18;   // Länge SEK Data
         LAENGE_VAL_DATA : Int := 8;   // Länge Value Data
         LAENGE_BIT_DATA : Int := 6;   // Länge Bit Data
         LAENGE_FKT : Int := 4;   // Länge Funktion
         Res16 : Int;   // Reserve
         Res18 : Int;   // Reserve
      END_STRUCT;
      SEK : Array[601..1000] of "UDT_SDC_EMS_TS_COM";   // Komando für Sektion
   END_VAR
BEGIN
END_DATA_BLOCK

DATA_BLOCK "DB_SDC_TS_IF_STATUS"   // DB3718
{ S7_Optimized_Access := 'FALSE' }
AUTHOR : FFM
FAMILY : SDC
NAME : SECT_IF